HMI tags "DB_SDC_POSITION_INSERTS"
   "DB_SDC_BARCODE_INSERTS_INSERT[19].COURSELOW" : DInt = PLC DB_SDC_BARCODE_INSERTS.INSERT[19].COURSELOW AT %DB3734.DBD364, 1 s   // lower position value Course Barocdevalue befor Insert
   "DB_SDC_BARCODE_INSERTS_INSERT[4].COURSEHIGH" : DInt = PLC DB_SDC_BARCODE_INSERTS.INSERT[4].COURSEHIGH AT %DB3734.DBD68, 1 s   // höhere Positionswert Course Barocde Wert nach Insert / higher position value Course Barocdevalue after Insert
   "DB_SDC_BARCODE_INSERTS_INSERT[15].INSERTHIGH" : DInt = PLC DB_SDC_BARCODE_INSERTS.INSERT[15].INSERTHIGH AT %DB3734.DBD296, 1 s   // höhere Positionswert Barocde Wert liegt Hoch / higher position value Barocdevalue Insert high
   "DB_SDC_BARCODE_INSERTS_INSERT[8].COURSELOW" : DInt = PLC DB_SDC_BARCODE_INSERTS.INSERT[8].COURSELOW AT %DB3734.DBD144, 1 s   // lower position value Course Barocdevalue befor Insert
   "DB_SDC_BARCODE_INSERTS_INSERT[9].INSERTLOW" : DInt = PLC DB_SDC_BARCODE_INSERTS.INSERT[9].INSERTLOW AT %DB3734.DBD172, 1 s   // lower position value Barocdevalue Insert low
   "DB_SDC_BARCODE_INSERTS_INSERT[14].COURSELOW" : DInt = PLC DB_SDC_BARCODE_INSERTS.INSERT[14].COURSELOW AT %DB3734.DBD264, 1 s   // lower position value Course Barocdevalue befor Insert
   "DB_SDC_BARCODE_INSERTS_INSERT[15].COURSEHIGH" : DInt = PLC DB_SDC_BARCODE_INSERTS.INSERT[15].COURSEHIGH AT %DB3734.DBD288, 1 s   // höhere Positionswert Course Barocde Wert nach Insert / higher position value Course Barocdevalue after Insert
   "DB_SDC_BARCODE_INSERTS_INSERT[19].COURSEHIGH" : DInt = PLC DB_SDC_BARCODE_INSERTS.INSERT[19].COURSEHIGH AT %DB3734.DBD368, 1 s   // höhere Positionswert Course Barocde Wert nach Insert / higher position value Course Barocdevalue after Insert
   "DB_SDC_BARCODE_INSERTS_INSERT[17].INSERTLOW" : DInt = PLC DB_SDC_BARCODE_INSERTS.INSERT[17].INSERTLOW AT %DB3734.DBD332, 1 s   // lower position value Barocdevalue Insert low
   "DB_SDC_BARCODE_INSERTS_INSERT[16].COURSEHIGH" : DInt = PLC DB_SDC_BARCODE_INSERTS.INSERT[16].COURSEHIGH AT %DB3734.DBD308, 1 s   // höhere Positionswert Course Barocde Wert nach Insert / higher position value Course Barocdevalue after Insert
   "DB_SDC_BARCODE_INSERTS_HYST" : Int = PLC DB_SDC_BARCODE_INSERTS.HYST AT %DB3734.DBW0, 1 s   // Hysterese für Positionswerte
   "DB_SDC_BARCODE_INSERTS_INSERT[3].OFFSET" : DInt = PLC DB_SDC_BARCODE_INSERTS.INSERT[3].OFFSET AT %DB3734.DBD60, 1 s   // absoluten Offset zu Beginn der Einfügen -> zusätzlich von allen Einsätzen unter / absolute offset at the start of the Insert -> addition from all inserts below
   "DB_SDC_BARCODE_INSERTS_INSERT[16].OFFSET" : DInt = PLC DB_SDC_BARCODE_INSERTS.INSERT[16].OFFSET AT %DB3734.DBD320, 1 s   // absoluten Offset zu Beginn der Einfügen -> zusätzlich von allen Einsätzen unter / absolute offset at the start of the Insert -> addition from all inserts below
   "DB_SDC_BARCODE_INSERTS_INSERT[10].OFFSET" : DInt = PLC DB_SDC_BARCODE_INSERTS.INSERT[10].OFFSET AT %DB3734.DBD200, 1 s   // absoluten Offset zu Beginn der Einfügen -> zusätzlich von allen Einsätzen unter / absolute offset at the start of the Insert -> addition from all inserts below
   "DB_SDC_BARCODE_INSERTS_INSERT[17].COURSELOW" : DInt = PLC DB_SDC_BARCODE_INSERTS.INSERT[17].COURSELOW AT %DB3734.DBD324, 1 s   // lower position value Course Barocdevalue befor Insert
   "DB_SDC_BARCODE_INSERTS_INSERT[4].INSERTLOW" : DInt = PLC DB_SDC_BARCODE_INSERTS.INSERT[4].INSERTLOW AT %DB3734.DBD72, 1 s   // lower position value Barocdevalue Insert low
   "DB_SDC_BARCODE_INSERTS_INSERT[20].COURSELOW" : DInt = PLC DB_SDC_BARCODE_INSERTS.INSERT[20].COURSELOW AT %DB3734.DBD384, 1 s   // lower position value Course Barocdevalue befor Insert
   "DB_SDC_BARCODE_INSERTS_INSERT[12].COURSELOW" : DInt = PLC DB_SDC_BARCODE_INSERTS.INSERT[12].COURSELOW AT %DB3734.DBD224, 1 s   // lower position value Course Barocdevalue befor Insert
   "DB_SDC_BARCODE_INSERTS_INSERT[7].COURSELOW" : DInt = PLC DB_SDC_BARCODE_INSERTS.INSERT[7].COURSELOW AT %DB3734.DBD124, 1 s   // lower position value Course Barocdevalue befor Insert
   "DB_SDC_BARCODE_INSERTS_INSERT[10].COURSELOW" : DInt = PLC DB_SDC_BARCODE_INSERTS.INSERT[10].COURSELOW AT %DB3734.DBD184, 1 s   // lower position value Course Barocdevalue befor Insert
   "DB_SDC_BARCODE_INSERTS_INSERT[3].COURSELOW" : DInt = PLC DB_SDC_BARCODE_INSERTS.INSERT[3].COURSELOW AT %DB3734.DBD44, 1 s   // lower position value Course Barocdevalue befor Insert
   "DB_SDC_BARCODE_INSERTS_INSERT[11].COURSELOW" : DInt = PLC DB_SDC_BARCODE_INSERTS.INSERT[11].COURSELOW AT %DB3734.DBD204, 1 s   // lower position value Course Barocdevalue befor Insert
   "DB_SDC_BARCODE_INSERTS_INSERT[15].COURSELOW" : DInt = PLC DB_SDC_BARCODE_INSERTS.INSERT[15].COURSELOW AT %DB3734.DBD284, 1 s   // lower position value Course Barocdevalue befor Insert
   "DB_SDC_BARCODE_INSERTS_INSERT[11].INSERTHIGH" : DInt = PLC DB_SDC_BARCODE_INSERTS.INSERT[11].INSERTHIGH AT %DB3734.DBD216, 1 s   // höhere Positionswert Barocde Wert liegt Hoch / higher position value Barocdevalue Insert high
   "DB_SDC_BARCODE_INSERTS_INSERT[17].INSERTHIGH" : DInt = PLC DB_SDC_BARCODE_INSERTS.INSERT[17].INSERTHIGH AT %DB3734.DBD336, 1 s   // höhere Positionswert Barocde Wert liegt Hoch / higher position value Barocdevalue Insert high
   "DB_SDC_BARCODE_INSERTS_INSERT[1].COURSEHIGH" : DInt = PLC DB_SDC_BARCODE_INSERTS.INSERT[1].COURSEHIGH AT %DB3734.DBD8, 1 s   // höhere Positionswert Course Barocde Wert nach Insert / higher position value Course Barocdevalue after Insert
   "DB_SDC_BARCODE_INSERTS_INSERT[11].OFFSET" : DInt = PLC DB_SDC_BARCODE_INSERTS.INSERT[11].OFFSET AT %DB3734.DBD220, 1 s   // absoluten Offset zu Beginn der Einfügen -> zusätzlich von allen Einsätzen unter / absolute offset at the start of the Insert -> addition from all inserts below
   "DB_SDC_BARCODE_INSERTS_INSERT[7].INSERTLOW" : DInt = PLC DB_SDC_BARCODE_INSERTS.INSERT[7].INSERTLOW AT %DB3734.DBD132, 1 s   // lower position value Barocdevalue Insert low
   "DB_SDC_BARCODE_INSERTS_INSERT[12].INSERTLOW" : DInt = PLC DB_SDC_BARCODE_INSERTS.INSERT[12].INSERTLOW AT %DB3734.DBD232, 1 s   // lower position value Barocdevalue Insert low
   "DB_SDC_BARCODE_INSERTS_INSERT[10].COURSEHIGH" : DInt = PLC DB_SDC_BARCODE_INSERTS.INSERT[10].COURSEHIGH AT %DB3734.DBD188, 1 s   // höhere Positionswert Course Barocde Wert nach Insert / higher position value Course Barocdevalue after Insert
   "DB_SDC_BARCODE_INSERTS_INSERTS" : Int = PLC DB_SDC_BARCODE_INSERTS.INSERTS AT %DB3734.DBW2, 1 s   // Positioning Leaps
   "DB_SDC_BARCODE_INSERTS_INSERT[8].INSERTHIGH" : DInt = PLC DB_SDC_BARCODE_INSERTS.INSERT[8].INSERTHIGH AT %DB3734.DBD156, 1 s   // höhere Positionswert Barocde Wert liegt Hoch / higher position value Barocdevalue Insert high
   "DB_SDC_BARCODE_INSERTS_INSERT[18].COURSELOW" : DInt = PLC DB_SDC_BARCODE_INSERTS.INSERT[18].COURSELOW AT %DB3734.DBD344, 1 s   // lower position value Course Barocdevalue befor Insert
   "DB_SDC_BARCODE_INSERTS_INSERT[5].INSERTHIGH" : DInt = PLC DB_SDC_BARCODE_INSERTS.INSERT[5].INSERTHIGH AT %DB3734.DBD96, 1 s   // höhere Positionswert Barocde Wert liegt Hoch / higher position value Barocdevalue Insert high
   "DB_SDC_BARCODE_INSERTS_INSERT[16].INSERTLOW" : DInt = PLC DB_SDC_BARCODE_INSERTS.INSERT[16].INSERTLOW AT %DB3734.DBD312, 1 s   // lower position value Barocdevalue Insert low
   "DB_SDC_BARCODE_INSERTS_INSERT[19].INSERTHIGH" : DInt = PLC DB_SDC_BARCODE_INSERTS.INSERT[19].INSERTHIGH AT %DB3734.DBD376, 1 s   // höhere Positionswert Barocde Wert liegt Hoch / higher position value Barocdevalue Insert high
   "DB_SDC_BARCODE_INSERTS_INSERT[18].COURSEHIGH" : DInt = PLC DB_SDC_BARCODE_INSERTS.INSERT[18].COURSEHIGH AT %DB3734.DBD348, 1 s   // höhere Positionswert Course Barocde Wert nach Insert / higher position value Course Barocdevalue after Insert
   "DB_SDC_BARCODE_INSERTS_INSERT[19].OFFSET" : DInt = PLC DB_SDC_BARCODE_INSERTS.INSERT[19].OFFSET AT %DB3734.DBD380, 1 s   // absoluten Offset zu Beginn der Einfügen -> zusätzlich von allen Einsätzen unter / absolute offset at the start of the Insert -> addition from all inserts below
   "DB_SDC_BARCODE_INSERTS_INSERT[8].INSERTLOW" : DInt = PLC DB_SDC_BARCODE_INSERTS.INSERT[8].INSERTLOW AT %DB3734.DBD152, 1 s   // lower position value Barocdevalue Insert low
   "DB_SDC_BARCODE_INSERTS_ABS_DIST_COURSE" : DInt = PLC DB_SDC_BARCODE_INSERTS.ABS_DIST_COURSE AT %DB3734.DBD404, 1 s   // abslolute Entfernung / abslolute Distance Course
   "DB_SDC_BARCODE_INSERTS_INSERT[14].INSERTLOW" : DInt = PLC DB_SDC_BARCODE_INSERTS.INSERT[14].INSERTLOW AT %DB3734.DBD272, 1 s   // lower position value Barocdevalue Insert low
   "DB_SDC_BARCODE_INSERTS_INSERT[13].COURSEHIGH" : DInt = PLC DB_SDC_BARCODE_INSERTS.INSERT[13].COURSEHIGH AT %DB3734.DBD248, 1 s   // höhere Positionswert Course Barocde Wert nach Insert / higher position value Course Barocdevalue after Insert
   "DB_SDC_BARCODE_INSERTS_INSERT[14].INSERTHIGH" : DInt = PLC DB_SDC_BARCODE_INSERTS.INSERT[14].INSERTHIGH AT %DB3734.DBD276, 1 s   // höhere Positionswert Barocde Wert liegt Hoch / higher position value Barocdevalue Insert high
   "DB_SDC_BARCODE_INSERTS_INSERT[5].INSERTLOW" : DInt = PLC DB_SDC_BARCODE_INSERTS.INSERT[5].INSERTLOW AT %DB3734.DBD92, 1 s   // lower position value Barocdevalue Insert low
   "DB_SDC_BARCODE_INSERTS_INSERT[14].OFFSET" : DInt = PLC DB_SDC_BARCODE_INSERTS.INSERT[14].OFFSET AT %DB3734.DBD280, 1 s   // absoluten Offset zu Beginn der Einfügen -> zusätzlich von allen Einsätzen unter / absolute offset at the start of the Insert -> addition from all inserts below
   "DB_SDC_BARCODE_INSERTS_INSERT[13].COURSELOW" : DInt = PLC DB_SDC_BARCODE_INSERTS.INSERT[13].COURSELOW AT %DB3734.DBD244, 1 s   // lower position value Course Barocdevalue befor Insert
   "DB_SDC_BARCODE_INSERTS_INSERT[7].COURSEHIGH" : DInt = PLC DB_SDC_BARCODE_INSERTS.INSERT[7].COURSEHIGH AT %DB3734.DBD128, 1 s   // höhere Positionswert Course Barocde Wert nach Insert / higher position value Course Barocdevalue after Insert
   "DB_SDC_BARCODE_INSERTS_INSERT[12].COURSEHIGH" : DInt = PLC DB_SDC_BARCODE_INSERTS.INSERT[12].COURSEHIGH AT %DB3734.DBD228, 1 s   // höhere Positionswert Course Barocde Wert nach Insert / higher position value Course Barocdevalue after Insert
   "DB_SDC_BARCODE_INSERTS_INSERT[18].INSERTHIGH" : DInt = PLC DB_SDC_BARCODE_INSERTS.INSERT[18].INSERTHIGH AT %DB3734.DBD356, 1 s   // höhere Positionswert Barocde Wert liegt Hoch / higher position value Barocdevalue Insert high
   "DB_SDC_BARCODE_INSERTS_INSERT[1].OFFSET" : DInt = PLC DB_SDC_BARCODE_INSERTS.INSERT[1].OFFSET AT %DB3734.DBD20, 1 s   // absoluten Offset zu Beginn der Einfügen -> zusätzlich von allen Einsätzen unter / absolute offset at the start of the Insert -> addition from all inserts below
   "DB_SDC_BARCODE_INSERTS_INSERT[1].INSERTHIGH" : DInt = PLC DB_SDC_BARCODE_INSERTS.INSERT[1].INSERTHIGH AT %DB3734.DBD16, 1 s   // höhere Positionswert Barocde Wert liegt Hoch / higher position value Barocdevalue Insert high
   "DB_SDC_BARCODE_INSERTS_INSERT[1].COURSELOW" : DInt = PLC DB_SDC_BARCODE_INSERTS.INSERT[1].COURSELOW AT %DB3734.DBD4, 1 s   // lower position value Course Barocdevalue befor Insert
   "DB_SDC_BARCODE_INSERTS_INSERT[3].INSERTHIGH" : DInt = PLC DB_SDC_BARCODE_INSERTS.INSERT[3].INSERTHIGH AT %DB3734.DBD56, 1 s   // höhere Positionswert Barocde Wert liegt Hoch / higher position value Barocdevalue Insert high
   "DB_SDC_BARCODE_INSERTS_INSERT[8].COURSEHIGH" : DInt = PLC DB_SDC_BARCODE_INSERTS.INSERT[8].COURSEHIGH AT %DB3734.DBD148, 1 s   // höhere Positionswert Course Barocde Wert nach Insert / higher position value Course Barocdevalue after Insert
   "DB_SDC_BARCODE_INSERTS_INSERT[5].OFFSET" : DInt = PLC DB_SDC_BARCODE_INSERTS.INSERT[5].OFFSET AT %DB3734.DBD100, 1 s   // absoluten Offset zu Beginn der Einfügen -> zusätzlich von allen Einsätzen unter / absolute offset at the start of the Insert -> addition from all inserts below
   "DB_SDC_BARCODE_INSERTS_INSERT[9].COURSELOW" : DInt = PLC DB_SDC_BARCODE_INSERTS.INSERT[9].COURSELOW AT %DB3734.DBD164, 1 s   // lower position value Course Barocdevalue befor Insert
   "DB_SDC_BARCODE_INSERTS_INSERT[14].COURSEHIGH" : DInt = PLC DB_SDC_BARCODE_INSERTS.INSERT[14].COURSEHIGH AT %DB3734.DBD268, 1 s   // höhere Positionswert Course Barocde Wert nach Insert / higher position value Course Barocdevalue after Insert
   "DB_SDC_BARCODE_INSERTS_INSERT[2].OFFSET" : DInt = PLC DB_SDC_BARCODE_INSERTS.INSERT[2].OFFSET AT %DB3734.DBD40, 1 s   // absoluten Offset zu Beginn der Einfügen -> zusätzlich von allen Einsätzen unter / absolute offset at the start of the Insert -> addition from all inserts below
   "DB_SDC_BARCODE_INSERTS_INSERT[17].OFFSET" : DInt = PLC DB_SDC_BARCODE_INSERTS.INSERT[17].OFFSET AT %DB3734.DBD340, 1 s   // absoluten Offset zu Beginn der Einfügen -> zusätzlich von allen Einsätzen unter / absolute offset at the start of the Insert -> addition from all inserts below
   "DB_SDC_BARCODE_INSERTS_INSERT[2].COURSELOW" : DInt = PLC DB_SDC_BARCODE_INSERTS.INSERT[2].COURSELOW AT %DB3734.DBD24, 1 s   // lower position value Course Barocdevalue befor Insert
   "DB_SDC_BARCODE_INSERTS_INSERT[16].COURSELOW" : DInt = PLC DB_SDC_BARCODE_INSERTS.INSERT[16].COURSELOW AT %DB3734.DBD304, 1 s   // lower position value Course Barocdevalue befor Insert
   "DB_SDC_BARCODE_INSERTS_INSERT[13].INSERTHIGH" : DInt = PLC DB_SDC_BARCODE_INSERTS.INSERT[13].INSERTHIGH AT %DB3734.DBD256, 1 s   // höhere Positionswert Barocde Wert liegt Hoch / higher position value Barocdevalue Insert high
   "DB_SDC_BARCODE_INSERTS_INSERT[2].INSERTHIGH" : DInt = PLC DB_SDC_BARCODE_INSERTS.INSERT[2].INSERTHIGH AT %DB3734.DBD36, 1 s   // höhere Positionswert Barocde Wert liegt Hoch / higher position value Barocdevalue Insert high
   "DB_SDC_BARCODE_INSERTS_INSERT[11].INSERTLOW" : DInt = PLC DB_SDC_BARCODE_INSERTS.INSERT[11].INSERTLOW AT %DB3734.DBD212, 1 s   // lower position value Barocdevalue Insert low
   "DB_SDC_BARCODE_INSERTS_INSERT[16].INSERTHIGH" : DInt = PLC DB_SDC_BARCODE_INSERTS.INSERT[16].INSERTHIGH AT %DB3734.DBD316, 1 s   // höhere Positionswert Barocde Wert liegt Hoch / higher position value Barocdevalue Insert high
   "DB_SDC_BARCODE_INSERTS_INSERT[20].COURSEHIGH" : DInt = PLC DB_SDC_BARCODE_INSERTS.INSERT[20].COURSEHIGH AT %DB3734.DBD388, 1 s   // höhere Positionswert Course Barocde Wert nach Insert / higher position value Course Barocdevalue after Insert
   "DB_SDC_BARCODE_INSERTS_INSERT[2].COURSEHIGH" : DInt = PLC DB_SDC_BARCODE_INSERTS.INSERT[2].COURSEHIGH AT %DB3734.DBD28, 1 s   // höhere Positionswert Course Barocde Wert nach Insert / higher position value Course Barocdevalue after Insert
   "DB_SDC_BARCODE_INSERTS_INSERT[5].COURSEHIGH" : DInt = PLC DB_SDC_BARCODE_INSERTS.INSERT[5].COURSEHIGH AT %DB3734.DBD88, 1 s   // höhere Positionswert Course Barocde Wert nach Insert / higher position value Course Barocdevalue after Insert
   "DB_SDC_BARCODE_INSERTS_INSERT[18].INSERTLOW" : DInt = PLC DB_SDC_BARCODE_INSERTS.INSERT[18].INSERTLOW AT %DB3734.DBD352, 1 s   // lower position value Barocdevalue Insert low
   "DB_SDC_BARCODE_INSERTS_INSERT[20].INSERTHIGH" : DInt = PLC DB_SDC_BARCODE_INSERTS.INSERT[20].INSERTHIGH AT %DB3734.DBD396, 1 s   // höhere Positionswert Barocde Wert liegt Hoch / higher position value Barocdevalue Insert high
   "DB_SDC_BARCODE_INSERTS_INSERT[15].OFFSET" : DInt = PLC DB_SDC_BARCODE_INSERTS.INSERT[15].OFFSET AT %DB3734.DBD300, 1 s   // absoluten Offset zu Beginn der Einfügen -> zusätzlich von allen Einsätzen unter / absolute offset at the start of the Insert -> addition from all inserts below
   "DB_SDC_BARCODE_INSERTS_INSERT[5].COURSELOW" : DInt = PLC DB_SDC_BARCODE_INSERTS.INSERT[5].COURSELOW AT %DB3734.DBD84, 1 s   // lower position value Course Barocdevalue befor Insert
   "DB_SDC_BARCODE_INSERTS_INSERT[2].INSERTLOW" : DInt = PLC DB_SDC_BARCODE_INSERTS.INSERT[2].INSERTLOW AT %DB3734.DBD32, 1 s   // lower position value Barocdevalue Insert low
   "DB_SDC_BARCODE_INSERTS_INSERT[12].OFFSET" : DInt = PLC DB_SDC_BARCODE_INSERTS.INSERT[12].OFFSET AT %DB3734.DBD240, 1 s   // absoluten Offset zu Beginn der Einfügen -> zusätzlich von allen Einsätzen unter / absolute offset at the start of the Insert -> addition from all inserts below
   "DB_SDC_BARCODE_INSERTS_INSERT[17].COURSEHIGH" : DInt = PLC DB_SDC_BARCODE_INSERTS.INSERT[17].COURSEHIGH AT %DB3734.DBD328, 1 s   // höhere Positionswert Course Barocde Wert nach Insert / higher position value Course Barocdevalue after Insert
   "DB_SDC_BARCODE_INSERTS_INSERT[4].INSERTHIGH" : DInt = PLC DB_SDC_BARCODE_INSERTS.INSERT[4].INSERTHIGH AT %DB3734.DBD76, 1 s   // höhere Positionswert Barocde Wert liegt Hoch / higher position value Barocdevalue Insert high
   "DB_SDC_BARCODE_INSERTS_INSERT[20].INSERTLOW" : DInt = PLC DB_SDC_BARCODE_INSERTS.INSERT[20].INSERTLOW AT %DB3734.DBD392, 1 s   // lower position value Barocdevalue Insert low
   "DB_SDC_BARCODE_INSERTS_INSERT[10].INSERTLOW" : DInt = PLC DB_SDC_BARCODE_INSERTS.INSERT[10].INSERTLOW AT %DB3734.DBD192, 1 s   // lower position value Barocdevalue Insert low
   "DB_SDC_BARCODE_INSERTS_INSERT[20].OFFSET" : DInt = PLC DB_SDC_BARCODE_INSERTS.INSERT[20].OFFSET AT %DB3734.DBD400, 1 s   // absoluten Offset zu Beginn der Einfügen -> zusätzlich von allen Einsätzen unter / absolute offset at the start of the Insert -> addition from all inserts below
   "DB_SDC_BARCODE_INSERTS_INSERT[4].COURSELOW" : DInt = PLC DB_SDC_BARCODE_INSERTS.INSERT[4].COURSELOW AT %DB3734.DBD64, 1 s   // lower position value Course Barocdevalue befor Insert
   "DB_SDC_BARCODE_INSERTS_INSERT[3].COURSEHIGH" : DInt = PLC DB_SDC_BARCODE_INSERTS.INSERT[3].COURSEHIGH AT %DB3734.DBD48, 1 s   // höhere Positionswert Course Barocde Wert nach Insert / higher position value Course Barocdevalue after Insert
   "DB_SDC_BARCODE_INSERTS_INSERT[6].COURSELOW" : DInt = PLC DB_SDC_BARCODE_INSERTS.INSERT[6].COURSELOW AT %DB3734.DBD104, 1 s   // lower position value Course Barocdevalue befor Insert
   "DB_SDC_BARCODE_INSERTS_INSERT[6].COURSEHIGH" : DInt = PLC DB_SDC_BARCODE_INSERTS.INSERT[6].COURSEHIGH AT %DB3734.DBD108, 1 s   // höhere Positionswert Course Barocde Wert nach Insert / higher position value Course Barocdevalue after Insert
   "DB_SDC_BARCODE_INSERTS_INSERT[3].INSERTLOW" : DInt = PLC DB_SDC_BARCODE_INSERTS.INSERT[3].INSERTLOW AT %DB3734.DBD52, 1 s   // lower position value Barocdevalue Insert low
   "DB_SDC_BARCODE_INSERTS_INSERT[12].INSERTHIGH" : DInt = PLC DB_SDC_BARCODE_INSERTS.INSERT[12].INSERTHIGH AT %DB3734.DBD236, 1 s   // höhere Positionswert Barocde Wert liegt Hoch / higher position value Barocdevalue Insert high
   "DB_SDC_BARCODE_INSERTS_INSERT[9].OFFSET" : DInt = PLC DB_SDC_BARCODE_INSERTS.INSERT[9].OFFSET AT %DB3734.DBD180, 1 s   // absoluten Offset zu Beginn der Einfügen -> zusätzlich von allen Einsätzen unter / absolute offset at the start of the Insert -> addition from all inserts below
   "DB_SDC_BARCODE_INSERTS_INSERT[9].COURSEHIGH" : DInt = PLC DB_SDC_BARCODE_INSERTS.INSERT[9].COURSEHIGH AT %DB3734.DBD168, 1 s   // höhere Positionswert Course Barocde Wert nach Insert / higher position value Course Barocdevalue after Insert
   "DB_SDC_BARCODE_INSERTS_INSERT[6].INSERTHIGH" : DInt = PLC DB_SDC_BARCODE_INSERTS.INSERT[6].INSERTHIGH AT %DB3734.DBD116, 1 s   // höhere Positionswert Barocde Wert liegt Hoch / higher position value Barocdevalue Insert high
   "DB_SDC_BARCODE_INSERTS_INSERT[6].INSERTLOW" : DInt = PLC DB_SDC_BARCODE_INSERTS.INSERT[6].INSERTLOW AT %DB3734.DBD112, 1 s   // lower position value Barocdevalue Insert low
   "DB_SDC_BARCODE_INSERTS_INSERT[7].INSERTHIGH" : DInt = PLC DB_SDC_BARCODE_INSERTS.INSERT[7].INSERTHIGH AT %DB3734.DBD136, 1 s   // höhere Positionswert Barocde Wert liegt Hoch / higher position value Barocdevalue Insert high
   "DB_SDC_BARCODE_INSERTS_INSERT[15].INSERTLOW" : DInt = PLC DB_SDC_BARCODE_INSERTS.INSERT[15].INSERTLOW AT %DB3734.DBD292, 1 s   // lower position value Barocdevalue Insert low
   "DB_SDC_BARCODE_INSERTS_INSERT[4].OFFSET" : DInt = PLC DB_SDC_BARCODE_INSERTS.INSERT[4].OFFSET AT %DB3734.DBD80, 1 s   // absoluten Offset zu Beginn der Einfügen -> zusätzlich von allen Einsätzen unter / absolute offset at the start of the Insert -> addition from all inserts below
   "DB_SDC_BARCODE_INSERTS_INSERT[9].INSERTHIGH" : DInt = PLC DB_SDC_BARCODE_INSERTS.INSERT[9].INSERTHIGH AT %DB3734.DBD176, 1 s   // höhere Positionswert Barocde Wert liegt Hoch / higher position value Barocdevalue Insert high
   "DB_SDC_BARCODE_INSERTS_INSERT[6].OFFSET" : DInt = PLC DB_SDC_BARCODE_INSERTS.INSERT[6].OFFSET AT %DB3734.DBD120, 1 s   // absoluten Offset zu Beginn der Einfügen -> zusätzlich von allen Einsätzen unter / absolute offset at the start of the Insert -> addition from all inserts below
   "DB_SDC_BARCODE_INSERTS_INSERT[13].INSERTLOW" : DInt = PLC DB_SDC_BARCODE_INSERTS.INSERT[13].INSERTLOW AT %DB3734.DBD252, 1 s   // lower position value Barocdevalue Insert low
   "DB_SDC_BARCODE_INSERTS_INSERT[19].INSERTLOW" : DInt = PLC DB_SDC_BARCODE_INSERTS.INSERT[19].INSERTLOW AT %DB3734.DBD372, 1 s   // lower position value Barocdevalue Insert low
   "DB_SDC_BARCODE_INSERTS_INSERT[11].COURSEHIGH" : DInt = PLC DB_SDC_BARCODE_INSERTS.INSERT[11].COURSEHIGH AT %DB3734.DBD208, 1 s   // höhere Positionswert Course Barocde Wert nach Insert / higher position value Course Barocdevalue after Insert
   "DB_SDC_BARCODE_INSERTS_INSERT[8].OFFSET" : DInt = PLC DB_SDC_BARCODE_INSERTS.INSERT[8].OFFSET AT %DB3734.DBD160, 1 s   // absoluten Offset zu Beginn der Einfügen -> zusätzlich von allen Einsätzen unter / absolute offset at the start of the Insert -> addition from all inserts below
   "DB_SDC_BARCODE_INSERTS_INSERT[13].OFFSET" : DInt = PLC DB_SDC_BARCODE_INSERTS.INSERT[13].OFFSET AT %DB3734.DBD260, 1 s   // absoluten Offset zu Beginn der Einfügen -> zusätzlich von allen Einsätzen unter / absolute offset at the start of the Insert -> addition from all inserts below
   "DB_SDC_BARCODE_INSERTS_INSERT[7].OFFSET" : DInt = PLC DB_SDC_BARCODE_INSERTS.INSERT[7].OFFSET AT %DB3734.DBD140, 1 s   // absoluten Offset zu Beginn der Einfügen -> zusätzlich von allen Einsätzen unter / absolute offset at the start of the Insert -> addition from all inserts below
   "DB_SDC_BARCODE_INSERTS_INSERT[10].INSERTHIGH" : DInt = PLC DB_SDC_BARCODE_INSERTS.INSERT[10].INSERTHIGH AT %DB3734.DBD196, 1 s   // höhere Positionswert Barocde Wert liegt Hoch / higher position value Barocdevalue Insert high
   "DB_SDC_BARCODE_INSERTS_INSERT[1].INSERTLOW" : DInt = PLC DB_SDC_BARCODE_INSERTS.INSERT[1].INSERTLOW AT %DB3734.DBD12, 1 s   // lower position value Barocdevalue Insert low
   "DB_SDC_BARCODE_INSERTS_INSERT[18].OFFSET" : DInt = PLC DB_SDC_BARCODE_INSERTS.INSERT[18].OFFSET AT %DB3734.DBD360, 1 s   // absoluten Offset zu Beginn der Einfügen -> zusätzlich von allen Einsätzen unter / absolute offset at the start of the Insert -> addition from all inserts below

HMI tags "DB_SDC_EMS_INFO"
   "EMS_Zone[1]" : UDT_ZoneStructure = PLC EMS.Zone[1] AT %DB8.DBX1034.0, 1 s
   "EMS_Zone[2]" : UDT_ZoneStructure = PLC EMS.Zone[2] AT %DB8.DBX2068.0, 1 s
   "EMS_Zone[3]" : UDT_ZoneStructure = PLC EMS.Zone[3] AT %DB8.DBX3102.0, 1 s
   "EMS_Zone[7]" : UDT_ZoneStructure = PLC EMS.Zone[7] AT %DB8.DBX7238.0, 1 s
   "EMS_Zone[8]" : UDT_ZoneStructure = PLC EMS.Zone[8] AT %DB8.DBX8272.0, 1 s
   "EMS_Zone[9]" : UDT_ZoneStructure = PLC EMS.Zone[9] AT %DB8.DBX9306.0, 1 s
   "EMS_Zone[10]" : UDT_ZoneStructure = PLC EMS.Zone[10] AT %DB8.DBX10340.0, 1 s
   "EMS_Zone[11]" : UDT_ZoneStructure = PLC EMS.Zone[11] AT %DB8.DBX11374.0, 1 s
   "EMS_Zone[12]" : UDT_ZoneStructure = PLC EMS.Zone[12] AT %DB8.DBX12408.0, 1 s
   "EMS_Zone[13]" : UDT_ZoneStructure = PLC EMS.Zone[13] AT %DB8.DBX13442.0, 1 s
   "EMS_Zone[14]" : UDT_ZoneStructure = PLC EMS.Zone[14] AT %DB8.DBX14476.0, 1 s
   "EMS_Zone[15]" : UDT_ZoneStructure = PLC EMS.Zone[15] AT %DB8.DBX15510.0, 1 s
   "EMS_Zone[16]" : UDT_ZoneStructure = PLC EMS.Zone[16] AT %DB8.DBX16544.0, 1 s
   "EMS_Zone[17]" : UDT_ZoneStructure = PLC EMS.Zone[17] AT %DB8.DBX17578.0, 1 s
   "EMS_Zone[18]" : UDT_ZoneStructure = PLC EMS.Zone[18] AT %DB8.DBX18612.0, 1 s
   "EMS_Zone[19]" : UDT_ZoneStructure = PLC EMS.Zone[19] AT %DB8.DBX19646.0, 1 s
   "EMS_Zone[20]" : UDT_ZoneStructure = PLC EMS.Zone[20] AT %DB8.DBX20680.0, 1 s
   "EMS_Zone[21]" : UDT_ZoneStructure = PLC EMS.Zone[21] AT %DB8.DBX21714.0, 1 s
   "EMS_Zone[22]" : UDT_ZoneStructure = PLC EMS.Zone[22] AT %DB8.DBX22748.0, 1 s
   "EMS_Zone[23]" : UDT_ZoneStructure = PLC EMS.Zone[23] AT %DB8.DBX23782.0, 1 s
   "EMS_Zone[24]" : UDT_ZoneStructure = PLC EMS.Zone[24] AT %DB8.DBX24816.0, 1 s
   "EMS_Zone[25]" : UDT_ZoneStructure = PLC EMS.Zone[25] AT %DB8.DBX25850.0, 1 s
   "EMS_Zone[26]" : UDT_ZoneStructure = PLC EMS.Zone[26] AT %DB8.DBX26884.0, 1 s
   "EMS_Zone[27]" : UDT_ZoneStructure = PLC EMS.Zone[27] AT %DB8.DBX27918.0, 1 s
   "EMS_Zone[28]" : UDT_ZoneStructure = PLC EMS.Zone[28] AT %DB8.DBX28952.0, 1 s
   "EMS_Zone[29]" : UDT_ZoneStructure = PLC EMS.Zone[29] AT %DB8.DBX29986.0, 1 s
   "EMS_Zone[30]" : UDT_ZoneStructure = PLC EMS.Zone[30] AT %DB8.DBX31020.0, 1 s
   "EMS_Carrier[1]" : UDT_CarrierStructure = PLC EMS.Carrier[1] AT %DB8.DBX63156.0, 1 s
   "EMS_Carrier[2]" : UDT_CarrierStructure = PLC EMS.Carrier[2] AT %DB8.DBX63238.0, 1 s
   "EMS_Carrier[3]" : UDT_CarrierStructure = PLC EMS.Carrier[3] AT %DB8.DBX63320.0, 1 s
   "EMS_Carrier[4]" : UDT_CarrierStructure = PLC EMS.Carrier[4] AT %DB8.DBX63402.0, 1 s
   "EMS_Carrier[5]" : UDT_CarrierStructure = PLC EMS.Carrier[5] AT %DB8.DBX63484.0, 1 s
   "EMS_Carrier[6]" : UDT_CarrierStructure = PLC EMS.Carrier[6] AT %DB8.DBX63566.0, 1 s
   "EMS_Carrier[7]" : UDT_CarrierStructure = PLC EMS.Carrier[7] AT %DB8.DBX63648.0, 1 s
   "EMS_Carrier[8]" : UDT_CarrierStructure = PLC EMS.Carrier[8] AT %DB8.DBX63730.0, 1 s
   "EMS_Carrier[9]" : UDT_CarrierStructure = PLC EMS.Carrier[9] AT %DB8.DBX63812.0, 1 s
   "EMS_Carrier[10]" : UDT_CarrierStructure = PLC DB_SDC_ERRORS_STAT.ER_AKT[42].ER_STAT[3].DRIVE_POS AT %DB8.DBX63894.0, 1 s
   "EMS_Carrier[11]" : UDT_CarrierStructure = PLC EMS.Carrier[11] AT %DB8.DBX63976.0, 1 s
   "EMS_Carrier[12]" : UDT_CarrierStructure = PLC EMS.Carrier[12] AT %DB8.DBX64058.0, 1 s
   "EMS_Carrier[13]" : UDT_CarrierStructure = PLC EMS.Carrier[13] AT %DB8.DBX64140.0, 1 s
   "EMS_Carrier[14]" : UDT_CarrierStructure = PLC EMS.Carrier[14] AT %DB8.DBX64222.0, 1 s
   "EMS_Carrier[15]" : UDT_CarrierStructure = PLC EMS.Carrier[15] AT %DB8.DBX64304.0, 1 s
   "EMS_Carrier[16]" : UDT_CarrierStructure = PLC EMS.Carrier[16] AT %DB8.DBX64386.0, 1 s
   "EMS_Carrier[17]" : UDT_CarrierStructure = PLC EMS.Carrier[17] AT %DB8.DBX64468.0, 1 s
   "EMS_Carrier[18]" : UDT_CarrierStructure = PLC EMS.Carrier[18] AT %DB8.DBX64550.0, 1 s
   "EMS_Carrier[19]" : UDT_CarrierStructure = PLC EMS.Carrier[19] AT %DB8.DBX64632.0, 1 s
   "EMS_Carrier[20]" : UDT_CarrierStructure = PLC EMS.Carrier[20] AT %DB8.DBX64714.0, 1 s
   "EMS_Carrier[21]" : UDT_CarrierStructure = PLC EMS.Carrier[21] AT %DB8.DBX64796.0, 1 s
   "EMS_Carrier[22]" : UDT_CarrierStructure = PLC EMS.Carrier[22] AT %DB8.DBX64878.0, 1 s
   "EMS_Carrier[23]" : UDT_CarrierStructure = PLC EMS.Carrier[23] AT %DB8.DBX64960.0, 1 s
   "EMS_Carrier[24]" : UDT_CarrierStructure = PLC EMS.Carrier[24] AT %DB8.DBX65042.0, 1 s
   "EMS_Carrier[25]" : UDT_CarrierStructure = PLC EMS.Carrier[25] AT %DB8.DBX65124.0, 1 s
   "EMS_Carrier[26]" : UDT_CarrierStructure = PLC EMS.Carrier[26] AT %DB8.DBX65206.0, 1 s
   "EMS_Carrier[27]" : UDT_CarrierStructure = PLC EMS.Carrier[27] AT %DB8.DBX65288.0, 1 s
   "EMS_Carrier[28]" : UDT_CarrierStructure = PLC EMS.Carrier[28] AT %DB8.DBX65370.0, 1 s
   "EMS_Carrier[29]" : UDT_CarrierStructure = PLC EMS.Carrier[29] AT %DB8.DBX65452.0, 1 s
   "EMS_Carrier[30]" : UDT_CarrierStructure = PLC EMS.Carrier[30], 1 s
   "EMS_Carrier[31]" : UDT_CarrierStructure = PLC EMS.Carrier[31], 1 s
   "EMS_Carrier[32]" : UDT_CarrierStructure = PLC EMS.Carrier[32], 1 s
   "EMS_Carrier[33]" : UDT_CarrierStructure = PLC EMS.Carrier[33], 1 s
   "EMS_Carrier[34]" : UDT_CarrierStructure = PLC EMS.Carrier[34], 1 s
   "EMS_Carrier[35]" : UDT_CarrierStructure = PLC EMS.Carrier[35], 1 s
   "EMS_Carrier[36]" : UDT_CarrierStructure = PLC EMS.Carrier[36], 1 s
   "EMS_Carrier[37]" : UDT_CarrierStructure = PLC EMS.Carrier[37], 1 s
   "EMS_Carrier[38]" : UDT_CarrierStructure = PLC EMS.Carrier[38], 1 s
   "EMS_Carrier[39]" : UDT_CarrierStructure = PLC EMS.Carrier[39], 1 s
   "EMS_Carrier[40]" : UDT_CarrierStructure = PLC EMS.Carrier[40], 1 s

HMI tags "DB_SDC_ERROR_STAT"
   "SDC\DB_SDC_ERROR_STAT\_Byte_DB_SDC_ERROR_STAT.F_STAT[XX5].EMS_TS_STAT_VAL.ERROR" : Int, internal   // Fehlernummer / Error number
   "SDC\DB_SDC_ERROR_STAT\_Byte_DB_SDC_ERROR_STAT.F_STAT[XX8].F" : Int, internal   // Fehler SDC + EMS Zusammenfassung / Fault SDC + EMS Summary
   "SDC\DB_SDC_ERROR_STAT\_Byte_DB_SDC_ERROR_STAT.F_STAT[X10].EMS_TS_STAT_VAL.DRIVE_POS_PERC" : Int, internal   // Position [% of Start End Section]
   "SDC\DB_SDC_ERROR_STAT\_Byte_DB_SDC_ERROR_STAT.F_STAT[XX9].F" : Int, internal   // Fehler SDC + EMS Zusammenfassung / Fault SDC + EMS Summary
   "SDC\DB_SDC_ERROR_STAT\_Byte_DB_SDC_ERROR_STAT.F_STAT[XX6].F_DATE" : Int, internal   // Fehler Zeit / Fault Time
   "SDC\DB_SDC_ERROR_STAT\DB_SDC_ERROR_STAT.F_STAT[XX7].EMS_TS_STAT_VAL.DRIVE_POS" : DInt AT %DB0.DBD0, 1 s   // Antriebsposition in mm / Drive position in mm
   "DB_SDC_ERRORS_STAT_HEADER.FAULT_PRO_SEITE_HMI" : Int = PLC DB_SDC_ERRORS_STAT.HEADER.FAULT_PRO_SEITE_HMI AT %DB3724.DBW10, 1 s   // Reserve
   "SDC\DB_SDC_ERROR_STAT\DB_SDC_ERROR_STAT.F_STAT[XX8].EMS_TS_STAT_VAL.DRIVE_POS" : DInt AT %DB0.DBD0, 1 s   // Antriebsposition in mm / Drive position in mm
   "SDC\DB_SDC_ERROR_STAT\DB_SDC_ERROR_STAT.F_STAT[XX8].EMS_TS_STAT_VAL.SEK" : Int AT %DB0.DBW0, 1 s   // Sektion
   "SDC\DB_SDC_ERROR_STAT\_Byte_DB_SDC_ERROR_STAT.F_STAT[XX1].EMS_TS_STAT_VAL.EMS_ID" : Int, internal   // EMS ID Nummer / EMS ID Number
   "SDC\DB_SDC_ERROR_STAT\DB_SDC_ERROR_STAT.F_STAT[XX5].EMS_TS_STAT_VAL.DRIVE_POS" : DInt AT %DB0.DBD0, 1 s   // Antriebsposition in mm / Drive position in mm
   "SDC\DB_SDC_ERROR_STAT\DB_SDC_ERROR_STAT.F_STAT[XX3].F_DATE" : Date_And_Time AT %DB0.DBX0.0, 1 s   // Fehler Zeit / Fault Time
   "SDC\DB_SDC_ERROR_STAT\_Byte_DB_SDC_ERROR_STAT.F_STAT[XX9].EMS_TS_STAT_VAL.TILT_POS" : Int, internal   // Tilt angle in degrees
   "SDC\DB_SDC_ERROR_STAT\DB_SDC_ERROR_STAT.F_STAT[XX7].F_DATE" : Date_And_Time AT %DB0.DBX0.0, 1 s   // Fehler Zeit / Fault Time
   "SDC\DB_SDC_ERROR_STAT\DB_SDC_ERROR_STAT.F_STAT[XX1].F_DATE" : Date_And_Time AT %DB0.DBX0.0, 1 s   // Fehler Zeit / Fault Time
   "SDC\DB_SDC_ERROR_STAT\DB_SDC_ERROR_STAT.F_STAT[XX4].EMS_TS_STAT_VAL.DRIVE_POS_PERC" : Int AT %DB0.DBW0, 1 s   // Position [% of Start End Section]
   "SDC\DB_SDC_ERROR_STAT\_Byte_DB_SDC_ERROR_STAT.F_STAT[XX6].EMS_TS_STAT_VAL.SEK" : Int, internal   // Sektion
   "SDC\DB_SDC_ERROR_STAT\_Byte_DB_SDC_ERROR_STAT.F_STAT[XX5].EMS_TS_STAT_VAL.PROFIL" : Int, internal   // Profile
   "SDC\DB_SDC_ERROR_STAT\DB_SDC_ERROR_STAT.F_STAT[XX5].EMS_TS_STAT_VAL.SEK" : Int AT %DB0.DBW0, 1 s   // Sektion
   "SDC\DB_SDC_ERROR_STAT\DB_SDC_ERROR_STAT.F_STAT[XX6].EMS_TS_STAT_VAL.PROFIL" : Int AT %DB0.DBW0, 1 s   // Profile
   "SDC\DB_SDC_ERROR_STAT\_Byte_DB_SDC_ERROR_STAT.F_STAT[XX8].EMS_TS_STAT_VAL.EMS_ID" : Int, internal   // EMS ID Nummer / EMS ID Number
   "SDC\DB_SDC_ERROR_STAT\_Byte_DB_SDC_ERROR_STAT.F_STAT[XX6].F" : Int, internal   // Fehler SDC + EMS Zusammenfassung / Fault SDC + EMS Summary
   "SDC\DB_SDC_ERROR_STAT\_Byte_DB_SDC_ERROR_STAT.F_STAT[XX5].EMS_TS_STAT_VAL.TILT_POS" : Int, internal   // Tilt angle in degrees
   "SDC\DB_SDC_ERROR_STAT\_Byte_DB_SDC_ERROR_STAT.F_STAT[XX2].EMS_TS_STAT_VAL.SEK" : Int, internal   // Sektion
   "SDC\DB_SDC_ERROR_STAT\DB_SDC_ERROR_STAT.F_STAT[XX5].F" : Word AT %DB0.DBW0, 1 s   // Fehler SDC + EMS Zusammenfassung / Fault SDC + EMS Summary
   "SDC\DB_SDC_ERROR_STAT\_Byte_DB_SDC_ERROR_STAT.F_STAT[XX7].F_DATE" : Int, internal   // Fehler Zeit / Fault Time
   "SDC\DB_SDC_ERROR_STAT\_Byte_DB_SDC_ERROR_STAT.F_STAT[XX6].EMS_TS_STAT_VAL.HOIST_POS" : Int, internal   // Höhe in mm / Height in mm
   "SDC\DB_SDC_ERROR_STAT\DB_SDC_ERROR_STAT.F_STAT[XX9].EMS_TS_STAT_VAL.HOIST_POS" : Int AT %DB0.DBW0, 1 s   // Höhe in mm / Height in mm
   "SDC\DB_SDC_ERROR_STAT\_Byte_DB_SDC_ERROR_STAT.F_STAT[XX1].EMS_TS_STAT_VAL.HOIST_POS" : Int, internal   // Höhe in mm / Height in mm
   "SDC\DB_SDC_ERROR_STAT\_Byte_DB_SDC_ERROR_STAT.F_STAT[XX5].EMS_TS_STAT_VAL.DRIVE_POS_PERC" : Int, internal   // Position [% of Start End Section]
   "SDC\DB_SDC_ERROR_STAT\DB_SDC_ERROR_STAT.F_STAT[XX1].EMS_TS_STAT_VAL.ERROR" : Int AT %DB0.DBW0, 1 s   // Fehlernummer / Error number
   "SDC\DB_SDC_ERROR_STAT\DB_SDC_ERROR_STAT.F_STAT[XX9].EMS_TS_STAT_VAL.SEK" : Int AT %DB0.DBW0, 1 s   // Sektion
   "SDC\DB_SDC_ERROR_STAT\_Byte_DB_SDC_ERROR_STAT.F_STAT[XX4].EMS_TS_STAT_VAL.DRIVE_POS" : Int, internal   // Antriebsposition in mm / Drive position in mm
   "SDC\DB_SDC_ERROR_STAT\DB_SDC_ERROR_STAT.F_STAT[XX4].EMS_TS_STAT_VAL.SEK" : Int AT %DB0.DBW0, 1 s   // Sektion
   "SDC\DB_SDC_ERROR_STAT\_Byte_DB_SDC_ERROR_STAT.F_STAT[XX2].F_DATE" : Int, internal   // Fehler Zeit / Fault Time
   "SDC\DB_SDC_ERROR_STAT\DB_SDC_ERROR_STAT.F_STAT[X10].EMS_TS_STAT_VAL.DRIVE_POS" : DInt AT %DB0.DBD0, 1 s   // Antriebsposition in mm / Drive position in mm
   "SDC\DB_SDC_ERROR_STAT\DB_SDC_ERROR_STAT.F_STAT[XX2].EMS_TS_STAT_VAL.TILT_POS" : Int AT %DB0.DBW0, 1 s   // Tilt angle in degrees
   "SDC\DB_SDC_ERROR_STAT\_Byte_DB_SDC_ERROR_STAT.F_STAT[XX2].EMS_TS_STAT_VAL.DRIVE_POS_PERC" : Int, internal   // Position [% of Start End Section]
   "SDC\DB_SDC_ERROR_STAT\_Byte_DB_SDC_ERROR_STAT.F_STAT[XX6].EMS_TS_STAT_VAL.TILT_POS" : Int, internal   // Tilt angle in degrees
   "SDC\DB_SDC_ERROR_STAT\DB_SDC_ERROR_STAT.F_STAT[XX5].EMS_TS_STAT_VAL.PROFIL" : Int AT %DB0.DBW0, 1 s   // Profile
   "SDC\DB_SDC_ERROR_STAT\_Byte_DB_SDC_ERROR_STAT.F_STAT[XX3].EMS_TS_STAT_VAL.EMS_ID" : Int, internal   // EMS ID Nummer / EMS ID Number
   "SDC\DB_SDC_ERROR_STAT\DB_SDC_ERROR_STAT.F_STAT[XX7].EMS_TS_STAT_VAL.SEK" : Int AT %DB0.DBW0, 1 s   // Sektion
   "SDC\DB_SDC_ERROR_STAT\DB_SDC_ERROR_STAT.F_STAT[XX1].EMS_TS_STAT_VAL.EMS_ID" : Int AT %DB0.DBW0, 1 s   // EMS ID Nummer / EMS ID Number
   "SDC\DB_SDC_ERROR_STAT\DB_SDC_ERROR_STAT.F_STAT[XX9].EMS_TS_STAT_VAL.TILT_POS" : Int AT %DB0.DBW0, 1 s   // Tilt angle in degrees
   "SDC\DB_SDC_ERROR_STAT\DB_SDC_ERROR_STAT.F_STAT[XX6].EMS_TS_STAT_VAL.HOIST_POS" : Int AT %DB0.DBW0, 1 s   // Höhe in mm / Height in mm
   "SDC\DB_SDC_ERROR_STAT\DB_SDC_ERROR_STAT.F_STAT[XX7].EMS_TS_STAT_VAL.PROFIL" : Int AT %DB0.DBW0, 1 s   // Profile